   Line "线_136#mig1_2" at 219,318 size 114x103
      Visibility <- "ST_HMI_Var_HMI_r64Axis_ChengXing_Position_real2"
   Line "线_3" at 219,227 size 125x91
      Visibility <- "ST_HMI_Var_HMI_r64Axis_ChengXing_Position_real2"
   Line "线_4" at 219,273 size 149x45
      Visibility <- "ST_HMI_Var_HMI_r64Axis_ChengXing_Position_real2"
   Line "线_11#mig1_2" at 219,225 size 124x93
      Visibility <- "ST_HMI_Var_HMI_r64Axis_ChengXing_Position_real2"
   Line "线_5" at 219,276 size 150x41
      Visibility <- "ST_HMI_Var_HMI_r64Axis_ChengXing_Position_real2"
   Line "线_6" at 219,318 size 112x105
      Visibility <- "ST_HMI_Var_HMI_r64Axis_ChengXing_Position_real2"
   Line "线_157" at 219,229 size 126x88
      Visibility <- "ST_HMI_Var_HMI_r64Axis_ChengXing_Position_real2"
   Line "线_115#mig1_2" at 219,318 size 155x11
      Visibility <- "ST_HMI_Var_HMI_r64Axis_ChengXing_Position_real2"
   Line "线_7" at 219,318 size 143x61
      Visibility <- "ST_HMI_Var_HMI_r64Axis_ChengXing_Position_real2"
   Line "线_159" at 219,318 size 155x13
      Visibility <- "ST_HMI_Var_HMI_r64Axis_ChengXing_Position_real2"
   Line "线_8" at 219,318 size 141x63
      Visibility <- "ST_HMI_Var_HMI_r64Axis_ChengXing_Position_real2"
   Line "线_9" at 219,318 size 110x106
      Visibility <- "ST_HMI_Var_HMI_r64Axis_ChengXing_Position_real2"
   Line "线_13#mig1_2" at 219,231 size 127x87
      Visibility <- "ST_HMI_Var_HMI_r64Axis_ChengXing_Position_real2"
   Line "线_14" at 219,278 size 151x39
      Visibility <- "ST_HMI_Var_HMI_r64Axis_ChengXing_Position_real2"
   Line "线_22" at 219,318 size 155x15
      Visibility <- "ST_HMI_Var_HMI_r64Axis_ChengXing_Position_real2"
   Line "线_24" at 219,318 size 140x66
      Visibility <- "ST_HMI_Var_HMI_r64Axis_ChengXing_Position_real2"
   Line "线_25" at 219,318 size 108x108
      Visibility <- "ST_HMI_Var_HMI_r64Axis_ChengXing_Position_real2"
   Line "线_124#mig1_2" at 219,234 size 129x84
      Visibility <- "ST_HMI_Var_HMI_r64Axis_ChengXing_Position_real2"
   Line "线_27" at 219,282 size 151x36
      Visibility <- "ST_HMI_Var_HMI_r64Axis_ChengXing_Position_real2"
   Line "线_195" at 219,318 size 155x18
      Visibility <- "ST_HMI_Var_HMI_r64Axis_ChengXing_Position_real2"
   Line "线_196" at 219,318 size 139x69
      Visibility <- "ST_HMI_Var_HMI_r64Axis_ChengXing_Position_real2"
   Line "线_197" at 219,318 size 106x111
      Visibility <- "ST_HMI_Var_HMI_r64Axis_ChengXing_Position_real2"
   Line "线_198" at 219,236 size 131x81
      Visibility <- "ST_HMI_Var_HMI_r64Axis_ChengXing_Position_real2"
   Line "线_199" at 219,284 size 151x33
      Visibility <- "ST_HMI_Var_HMI_r64Axis_ChengXing_Position_real2"
   Line "线_200" at 219,318 size 154x21
      Visibility <- "ST_HMI_Var_HMI_r64Axis_ChengXing_Position_real2"
   Line "线_201" at 219,318 size 138x70
      Visibility <- "ST_HMI_Var_HMI_r64Axis_ChengXing_Position_real2"
   Line "线_202" at 219,318 size 104x112
      Visibility <- "ST_HMI_Var_HMI_r64Axis_ChengXing_Position_real2"
   Line "线_254" at 219,238 size 132x80
      Visibility <- "ST_HMI_Var_HMI_r64Axis_ChengXing_Position_real2"
   Line "线_255" at 219,287 size 152x31
      Visibility <- "ST_HMI_Var_HMI_r64Axis_ChengXing_Position_real2"
   Line "线_256" at 219,318 size 154x23
      Visibility <- "ST_HMI_Var_HMI_r64Axis_ChengXing_Position_real2"
   Line "线_257" at 219,318 size 136x73
      Visibility <- "ST_HMI_Var_HMI_r64Axis_ChengXing_Position_real2"
   Line "线_277" at 219,318 size 102x114
      Visibility <- "ST_HMI_Var_HMI_r64Axis_ChengXing_Position_real2"
   Line "线_278" at 219,240 size 133x77
      Visibility <- "ST_HMI_Var_HMI_r64Axis_ChengXing_Position_real2"
   Line "线_279" at 219,289 size 153x28
      Visibility <- "ST_HMI_Var_HMI_r64Axis_ChengXing_Position_real2"
   Line "线_280" at 219,318 size 153x27
      Visibility <- "ST_HMI_Var_HMI_r64Axis_ChengXing_Position_real2"
   Line "线_281" at 219,318 size 135x75
      Visibility <- "ST_HMI_Var_HMI_r64Axis_ChengXing_Position_real2"
   Line "线_282" at 219,318 size 100x116
      Visibility <- "ST_HMI_Var_HMI_r64Axis_ChengXing_Position_real2"
   Line "线_283" at 219,243 size 135x75
      Visibility <- "ST_HMI_Var_HMI_r64Axis_ChengXing_Position_real2"
   Line "线_125#mig1_2" at 219,291 size 153x27
      Visibility <- "ST_HMI_Var_HMI_r64Axis_ChengXing_Position_real2"
   Line "线_284" at 219,318 size 153x28
      Visibility <- "ST_HMI_Var_HMI_r64Axis_ChengXing_Position_real2"
   Line "线_285" at 219,318 size 133x77
      Visibility <- "ST_HMI_Var_HMI_r64Axis_ChengXing_Position_real2"
   Line "线_286" at 219,318 size 98x117
      Visibility <- "ST_HMI_Var_HMI_r64Axis_ChengXing_Position_real2"
   Line "线_287" at 219,245 size 136x73
      Visibility <- "ST_HMI_Var_HMI_r64Axis_ChengXing_Position_real2"
   Line "线_288" at 219,294 size 154x24
      Visibility <- "ST_HMI_Var_HMI_r64Axis_ChengXing_Position_real2"
   Line "线_289" at 219,318 size 152x32
      Visibility <- "ST_HMI_Var_HMI_r64Axis_ChengXing_Position_real2"
   Line "线_290" at 219,318 size 132x80
      Visibility <- "ST_HMI_Var_HMI_r64Axis_ChengXing_Position_real2"
   Line "线_291" at 219,318 size 96x119
      Visibility <- "ST_HMI_Var_HMI_r64Axis_ChengXing_Position_real2"
   Line "线_292" at 219,246 size 138x71
      Visibility <- "ST_HMI_Var_HMI_r64Axis_ChengXing_Position_real2"
   Line "线_293" at 219,296 size 155x21
      Visibility <- "ST_HMI_Var_HMI_r64Axis_ChengXing_Position_real2"
   Line "线_294" at 219,318 size 151x33
      Visibility <- "ST_HMI_Var_HMI_r64Axis_ChengXing_Position_real2"
   Line "线_295" at 219,318 size 131x82
      Visibility <- "ST_HMI_Var_HMI_r64Axis_ChengXing_Position_real2"
   Line "线_315" at 219,318 size 93x121
      Visibility <- "ST_HMI_Var_HMI_r64Axis_ChengXing_Position_real2"
   Line "线_316" at 219,249 size 139x69
      Visibility <- "ST_HMI_Var_HMI_r64Axis_ChengXing_Position_real2"
   Line "线_130#mig1_2" at 219,299 size 155x19
      Visibility <- "ST_HMI_Var_HMI_r64Axis_ChengXing_Position_real2"
   Line "线_317" at 219,318 size 92x123
      Visibility <- "ST_HMI_Var_HMI_r64Axis_ChengXing_Position_real2"
   Line "线_97#mig1_2" at 219,251 size 140x67
      Visibility <- "ST_HMI_Var_HMI_r64Axis_ChengXing_Position_real2"
   Line "线_129#mig1_2" at 219,301 size 155x16
      Visibility <- "ST_HMI_Var_HMI_r64Axis_ChengXing_Position_real2"
   Line "线_318" at 219,318 size 151x37
      Visibility <- "ST_HMI_Var_HMI_r64Axis_ChengXing_Position_real2"
   Line "线_319" at 219,318 size 129x84
      Visibility <- "ST_HMI_Var_HMI_r64Axis_ChengXing_Position_real2"
   Line "线_320" at 219,318 size 89x123
      Visibility <- "ST_HMI_Var_HMI_r64Axis_ChengXing_Position_real2"
   Line "线_321" at 219,253 size 141x64
      Visibility <- "ST_HMI_Var_HMI_r64Axis_ChengXing_Position_real2"
   Line "线_128#mig1_2" at 219,305 size 155x13
      Visibility <- "ST_HMI_Var_HMI_r64Axis_ChengXing_Position_real2"
   Line "线_322" at 219,318 size 151x39
      Visibility <- "ST_HMI_Var_HMI_r64Axis_ChengXing_Position_real2"
   Line "线_323" at 219,318 size 127x87
      Visibility <- "ST_HMI_Var_HMI_r64Axis_ChengXing_Position_real2"
   Line "线_324" at 219,256 size 143x62
      Visibility <- "ST_HMI_Var_HMI_r64Axis_ChengXing_Position_real2"
   Line "线_131#mig1_2" at 219,306 size 155x11
      Visibility <- "ST_HMI_Var_HMI_r64Axis_ChengXing_Position_real2"
   Line "线_325" at 219,318 size 150x42
      Visibility <- "ST_HMI_Var_HMI_r64Axis_ChengXing_Position_real2"
   Line "线_326" at 219,318 size 126x89
      Visibility <- "ST_HMI_Var_HMI_r64Axis_ChengXing_Position_real2"
   Line "线_114#mig1_2" at 219,258 size 144x59
      Visibility <- "ST_HMI_Var_HMI_r64Axis_ChengXing_Position_real2"
   Line "线_327" at 219,310 size 156x8
      Visibility <- "ST_HMI_Var_HMI_r64Axis_ChengXing_Position_real2"
   Line "线_328" at 219,318 size 149x45
      Visibility <- "ST_HMI_Var_HMI_r64Axis_ChengXing_Position_real2"
   Line "线_329" at 219,318 size 125x91
      Visibility <- "ST_HMI_Var_HMI_r64Axis_ChengXing_Position_real2"
   Line "线_120#mig1_2" at 219,261 size 144x57
      Visibility <- "ST_HMI_Var_HMI_r64Axis_ChengXing_Position_real2"
   Line "线_330" at 219,312 size 156x5
      Visibility <- "ST_HMI_Var_HMI_r64Axis_ChengXing_Position_real2"
   Line "线_331" at 219,318 size 148x47
      Visibility <- "ST_HMI_Var_HMI_r64Axis_ChengXing_Position_real2"
   Line "线_332" at 219,318 size 123x93
      Visibility <- "ST_HMI_Var_HMI_r64Axis_ChengXing_Position_real2"
   Line "线_333" at 219,264 size 145x54
      Visibility <- "ST_HMI_Var_HMI_r64Axis_ChengXing_Position_real2"
   Line "线_150#mig1_2" at 219,315 size 156x3
      Visibility <- "ST_HMI_Var_HMI_r64Axis_ChengXing_Position_real2"
   Line "线_334" at 219,318 size 147x50
      Visibility <- "ST_HMI_Var_HMI_r64Axis_ChengXing_Position_real2"
   Line "线_335" at 219,318 size 121x95
      Visibility <- "ST_HMI_Var_HMI_r64Axis_ChengXing_Position_real2"
   Line "线_336" at 219,266 size 146x51
      Visibility <- "ST_HMI_Var_HMI_r64Axis_ChengXing_Position_real2"
   Line "线_147#mig1_2" at 219,318 size 156x0
      Visibility <- "ST_HMI_Var_HMI_r64Axis_ChengXing_Position_real2"
   Line "线_337" at 219,318 size 146x52
      Visibility <- "ST_HMI_Var_HMI_r64Axis_ChengXing_Position_real2"
   Line "线_338" at 219,318 size 119x98
      Visibility <- "ST_HMI_Var_HMI_r64Axis_ChengXing_Position_real2"
   Line "线_339" at 219,268 size 147x50
      Visibility <- "ST_HMI_Var_HMI_r64Axis_ChengXing_Position_real2"
   Line "线_340" at 219,318 size 156x3
      Visibility <- "ST_HMI_Var_HMI_r64Axis_ChengXing_Position_real2"
   Line "线_341" at 219,318 size 145x54
      Visibility <- "ST_HMI_Var_HMI_r64Axis_ChengXing_Position_real2"
   Line "线_342" at 219,318 size 144x57
      Visibility <- "ST_HMI_Var_HMI_r64Axis_ChengXing_Position_real2"
   Line "线_343" at 219,318 size 118x99
      Visibility <- "ST_HMI_Var_HMI_r64Axis_ChengXing_Position_real2"
   Line "线_344" at 219,318 size 116x101
      Visibility <- "ST_HMI_Var_HMI_r64Axis_ChengXing_Position_real2"
   Line "线_345" at 219,271 size 148x46
      Visibility <- "ST_HMI_Var_HMI_r64Axis_ChengXing_Position_real2"
   Line "线_346" at 219,318 size 156x5
      Visibility <- "ST_HMI_Var_HMI_r64Axis_ChengXing_Position_real2"
   Line "线_29" at 219,318 size 156x8
      Visibility <- "ST_HMI_Var_HMI_r64Axis_ChengXing_Position_real2"
   Line "线_31" at 219,318 size 144x58
      Visibility <- "ST_HMI_Var_HMI_r64Axis_ChengXing_Position_real2"
   Line "线_136#mig1_1" at 219,318 size 114x103
      Visibility <- "ST_HMI_Var_HMI_r64Axis_ChengXing_Position_real2"
   Line "线_38" at 219,227 size 125x91
      Visibility <- "ST_HMI_Var_HMI_r64Axis_ChengXing_Position_real2"
   Line "线_39" at 219,273 size 149x45
      Visibility <- "ST_HMI_Var_HMI_r64Axis_ChengXing_Position_real2"
   Line "线_11#mig1_1" at 219,225 size 124x93
      Visibility <- "ST_HMI_Var_HMI_r64Axis_ChengXing_Position_real2"
   Line "线_41" at 219,276 size 150x41
      Visibility <- "ST_HMI_Var_HMI_r64Axis_ChengXing_Position_real2"
   Line "线_43" at 219,318 size 112x105
      Visibility <- "ST_HMI_Var_HMI_r64Axis_ChengXing_Position_real2"
   Line "线_44" at 219,229 size 126x88
      Visibility <- "ST_HMI_Var_HMI_r64Axis_ChengXing_Position_real2"
   Line "线_115#mig1_1" at 219,318 size 155x11
      Visibility <- "ST_HMI_Var_HMI_r64Axis_ChengXing_Position_real2"
   Line "线_46" at 219,318 size 143x61
      Visibility <- "ST_HMI_Var_HMI_r64Axis_ChengXing_Position_real2"
   Line "线_47" at 219,318 size 155x13
      Visibility <- "ST_HMI_Var_HMI_r64Axis_ChengXing_Position_real2"
   Line "线_48" at 219,318 size 141x63
      Visibility <- "ST_HMI_Var_HMI_r64Axis_ChengXing_Position_real2"
   Line "线_49" at 219,318 size 110x106
      Visibility <- "ST_HMI_Var_HMI_r64Axis_ChengXing_Position_real2"
   Line "线_13#mig1_1" at 219,231 size 127x87
      Visibility <- "ST_HMI_Var_HMI_r64Axis_ChengXing_Position_real2"
   Line "线_59" at 219,278 size 151x39
      Visibility <- "ST_HMI_Var_HMI_r64Axis_ChengXing_Position_real2"
   Line "线_60" at 219,318 size 155x15
      Visibility <- "ST_HMI_Var_HMI_r64Axis_ChengXing_Position_real2"
   Line "线_61" at 219,318 size 140x66
      Visibility <- "ST_HMI_Var_HMI_r64Axis_ChengXing_Position_real2"
   Line "线_65" at 219,318 size 108x108
      Visibility <- "ST_HMI_Var_HMI_r64Axis_ChengXing_Position_real2"
   Line "线_124#mig1_1" at 219,234 size 129x84
      Visibility <- "ST_HMI_Var_HMI_r64Axis_ChengXing_Position_real2"
   Line "线_66" at 219,282 size 151x36
      Visibility <- "ST_HMI_Var_HMI_r64Axis_ChengXing_Position_real2"
   Line "线_67" at 219,318 size 155x18
      Visibility <- "ST_HMI_Var_HMI_r64Axis_ChengXing_Position_real2"
   Line "线_69" at 219,318 size 139x69
      Visibility <- "ST_HMI_Var_HMI_r64Axis_ChengXing_Position_real2"
   Line "线_70" at 219,318 size 106x111
      Visibility <- "ST_HMI_Var_HMI_r64Axis_ChengXing_Position_real2"
   Line "线_71" at 219,236 size 131x81
      Visibility <- "ST_HMI_Var_HMI_r64Axis_ChengXing_Position_real2"
   Line "线_72" at 219,284 size 151x33
      Visibility <- "ST_HMI_Var_HMI_r64Axis_ChengXing_Position_real2"
   Line "线_73" at 219,318 size 154x21
      Visibility <- "ST_HMI_Var_HMI_r64Axis_ChengXing_Position_real2"
   Line "线_74" at 219,318 size 138x70
      Visibility <- "ST_HMI_Var_HMI_r64Axis_ChengXing_Position_real2"
   Line "线_76" at 219,318 size 104x112
      Visibility <- "ST_HMI_Var_HMI_r64Axis_ChengXing_Position_real2"
   Line "线_77" at 219,238 size 132x80
      Visibility <- "ST_HMI_Var_HMI_r64Axis_ChengXing_Position_real2"
   Line "线_78" at 219,287 size 152x31
      Visibility <- "ST_HMI_Var_HMI_r64Axis_ChengXing_Position_real2"
   Line "线_79" at 219,318 size 154x23
      Visibility <- "ST_HMI_Var_HMI_r64Axis_ChengXing_Position_real2"
   Line "线_82" at 219,318 size 136x73
      Visibility <- "ST_HMI_Var_HMI_r64Axis_ChengXing_Position_real2"
   Line "线_84" at 219,318 size 102x114
      Visibility <- "ST_HMI_Var_HMI_r64Axis_ChengXing_Position_real2"
   Line "线_86" at 219,240 size 133x77
      Visibility <- "ST_HMI_Var_HMI_r64Axis_ChengXing_Position_real2"
   Line "线_87" at 219,289 size 153x28
      Visibility <- "ST_HMI_Var_HMI_r64Axis_ChengXing_Position_real2"
   Line "线_88" at 219,318 size 153x27
      Visibility <- "ST_HMI_Var_HMI_r64Axis_ChengXing_Position_real2"
   Line "线_90" at 219,318 size 135x75
      Visibility <- "ST_HMI_Var_HMI_r64Axis_ChengXing_Position_real2"
   Line "线_92" at 219,318 size 100x116
      Visibility <- "ST_HMI_Var_HMI_r64Axis_ChengXing_Position_real2"
   Line "线_93" at 219,243 size 135x75
      Visibility <- "ST_HMI_Var_HMI_r64Axis_ChengXing_Position_real2"
   Line "线_125#mig1_1" at 219,291 size 153x27
      Visibility <- "ST_HMI_Var_HMI_r64Axis_ChengXing_Position_real2"
   Line "线_98" at 219,318 size 153x28
      Visibility <- "ST_HMI_Var_HMI_r64Axis_ChengXing_Position_real2"
   Line "线_99" at 219,318 size 133x77
      Visibility <- "ST_HMI_Var_HMI_r64Axis_ChengXing_Position_real2"
   Line "线_109" at 219,318 size 98x117
      Visibility <- "ST_HMI_Var_HMI_r64Axis_ChengXing_Position_real2"
   Line "线_117" at 219,245 size 136x73
      Visibility <- "ST_HMI_Var_HMI_r64Axis_ChengXing_Position_real2"
   Line "线_119" at 219,294 size 154x24
      Visibility <- "ST_HMI_Var_HMI_r64Axis_ChengXing_Position_real2"
   Line "线_132" at 219,318 size 152x32
      Visibility <- "ST_HMI_Var_HMI_r64Axis_ChengXing_Position_real2"
   Line "线_135" at 219,318 size 132x80
      Visibility <- "ST_HMI_Var_HMI_r64Axis_ChengXing_Position_real2"
   Line "线_138" at 219,318 size 96x119
      Visibility <- "ST_HMI_Var_HMI_r64Axis_ChengXing_Position_real2"
   Line "线_347" at 219,246 size 138x71
      Visibility <- "ST_HMI_Var_HMI_r64Axis_ChengXing_Position_real2"
   Line "线_348" at 219,296 size 155x21
      Visibility <- "ST_HMI_Var_HMI_r64Axis_ChengXing_Position_real2"
   Line "线_349" at 219,318 size 151x33
      Visibility <- "ST_HMI_Var_HMI_r64Axis_ChengXing_Position_real2"
   Line "线_350" at 219,318 size 131x82
      Visibility <- "ST_HMI_Var_HMI_r64Axis_ChengXing_Position_real2"
   Line "线_351" at 219,318 size 93x121
      Visibility <- "ST_HMI_Var_HMI_r64Axis_ChengXing_Position_real2"
   Line "线_352" at 219,249 size 139x69
      Visibility <- "ST_HMI_Var_HMI_r64Axis_ChengXing_Position_real2"
   Line "线_130#mig1_1" at 219,299 size 155x19
      Visibility <- "ST_HMI_Var_HMI_r64Axis_ChengXing_Position_real2"
   Line "线_353" at 219,318 size 92x123
      Visibility <- "ST_HMI_Var_HMI_r64Axis_ChengXing_Position_real2"
   Line "线_97#mig1_1" at 219,251 size 140x67
      Visibility <- "ST_HMI_Var_HMI_r64Axis_ChengXing_Position_real2"
   Line "线_129#mig1_1" at 219,301 size 155x16
      Visibility <- "ST_HMI_Var_HMI_r64Axis_ChengXing_Position_real2"
   Line "线_354" at 219,318 size 151x37
      Visibility <- "ST_HMI_Var_HMI_r64Axis_ChengXing_Position_real2"
   Line "线_355" at 219,318 size 129x84
      Visibility <- "ST_HMI_Var_HMI_r64Axis_ChengXing_Position_real2"
   Line "线_356" at 219,318 size 89x123
      Visibility <- "ST_HMI_Var_HMI_r64Axis_ChengXing_Position_real2"
   Line "线_357" at 219,253 size 141x64
      Visibility <- "ST_HMI_Var_HMI_r64Axis_ChengXing_Position_real2"
   Line "线_128#mig1_1" at 219,305 size 155x13
      Visibility <- "ST_HMI_Var_HMI_r64Axis_ChengXing_Position_real2"
   Line "线_358" at 219,318 size 151x39
      Visibility <- "ST_HMI_Var_HMI_r64Axis_ChengXing_Position_real2"
   Line "线_359" at 219,318 size 127x87
      Visibility <- "ST_HMI_Var_HMI_r64Axis_ChengXing_Position_real2"
   Line "线_360" at 219,256 size 143x62
      Visibility <- "ST_HMI_Var_HMI_r64Axis_ChengXing_Position_real2"
   Line "线_131#mig1_1" at 219,306 size 155x11
      Visibility <- "ST_HMI_Var_HMI_r64Axis_ChengXing_Position_real2"
   Line "线_361" at 219,318 size 150x42
      Visibility <- "ST_HMI_Var_HMI_r64Axis_ChengXing_Position_real2"
   Line "线_362" at 219,318 size 126x89
      Visibility <- "ST_HMI_Var_HMI_r64Axis_ChengXing_Position_real2"
   Line "线_114#mig1_1" at 219,258 size 144x59
      Visibility <- "ST_HMI_Var_HMI_r64Axis_ChengXing_Position_real2"
   Line "线_363" at 219,310 size 156x8
      Visibility <- "ST_HMI_Var_HMI_r64Axis_ChengXing_Position_real2"
   Line "线_364" at 219,318 size 149x45
      Visibility <- "ST_HMI_Var_HMI_r64Axis_ChengXing_Position_real2"
   Line "线_365" at 219,318 size 125x91
      Visibility <- "ST_HMI_Var_HMI_r64Axis_ChengXing_Position_real2"
   Line "线_120#mig1_1" at 219,261 size 144x57
      Visibility <- "ST_HMI_Var_HMI_r64Axis_ChengXing_Position_real2"
   Line "线_366" at 219,312 size 156x5
      Visibility <- "ST_HMI_Var_HMI_r64Axis_ChengXing_Position_real2"
   Line "线_367" at 219,318 size 148x47
      Visibility <- "ST_HMI_Var_HMI_r64Axis_ChengXing_Position_real2"
   Line "线_368" at 219,318 size 123x93
      Visibility <- "ST_HMI_Var_HMI_r64Axis_ChengXing_Position_real2"
   Line "线_369" at 219,264 size 145x54
      Visibility <- "ST_HMI_Var_HMI_r64Axis_ChengXing_Position_real2"
   Line "线_150#mig1_1" at 219,315 size 156x3
      Visibility <- "ST_HMI_Var_HMI_r64Axis_ChengXing_Position_real2"
   Line "线_370" at 219,318 size 147x50
      Visibility <- "ST_HMI_Var_HMI_r64Axis_ChengXing_Position_real2"
   Line "线_371" at 219,318 size 121x95
      Visibility <- "ST_HMI_Var_HMI_r64Axis_ChengXing_Position_real2"
   Line "线_372" at 219,266 size 146x51
      Visibility <- "ST_HMI_Var_HMI_r64Axis_ChengXing_Position_real2"
   Line "线_147#mig1_1" at 219,318 size 156x0
      Visibility <- "ST_HMI_Var_HMI_r64Axis_ChengXing_Position_real2"
   Line "线_373" at 219,318 size 146x52
      Visibility <- "ST_HMI_Var_HMI_r64Axis_ChengXing_Position_real2"
   Line "线_374" at 219,318 size 119x98
      Visibility <- "ST_HMI_Var_HMI_r64Axis_ChengXing_Position_real2"
   Line "线_375" at 219,268 size 147x50
      Visibility <- "ST_HMI_Var_HMI_r64Axis_ChengXing_Position_real2"
   Line "线_376" at 219,318 size 156x3
      Visibility <- "ST_HMI_Var_HMI_r64Axis_ChengXing_Position_real2"
   Line "线_377" at 219,318 size 145x54
      Visibility <- "ST_HMI_Var_HMI_r64Axis_ChengXing_Position_real2"
   Line "线_378" at 219,318 size 144x57
      Visibility <- "ST_HMI_Var_HMI_r64Axis_ChengXing_Position_real2"
   Line "线_379" at 219,318 size 118x99
      Visibility <- "ST_HMI_Var_HMI_r64Axis_ChengXing_Position_real2"
   Line "线_380" at 219,318 size 116x101
      Visibility <- "ST_HMI_Var_HMI_r64Axis_ChengXing_Position_real2"
   Line "线_381" at 219,271 size 148x46
      Visibility <- "ST_HMI_Var_HMI_r64Axis_ChengXing_Position_real2"
   Line "线_382" at 219,318 size 156x5
      Visibility <- "ST_HMI_Var_HMI_r64Axis_ChengXing_Position_real2"
   Polygon "多边形_8" at 292,385 size 21x46
      Visibility <- "VBS_hengsi_status0"
   Polygon "多边形_7" at 288,376 size 31x55
      Visibility <- "VBS_hengsi_status0"
   Polygon "多边形_10" at 287,367 size 36x63
      Visibility <- "VBS_hengsi_status0"
   Polygon "多边形_11#mig1" at 287,361 size 40x70
      Visibility <- "VBS_hengsi_status0"
   Polygon "多边形_12" at 285,354 size 45x77
      Visibility <- "VBS_hengsi_status0"
   Polygon "多边形_18" at 285,345 size 45x86
      Visibility <- "VBS_hengsi_status1"
   Polygon "多边形_17" at 285,338 size 49x93
      Visibility <- "VBS_hengsi_status1"
   Polygon "多边形_16" at 287,328 size 50x103
      Visibility <- "VBS_hengsi_status1"
   Polygon "多边形_15" at 287,318 size 54x115
      Visibility <- "VBS_hengsi_status1"
   Polygon "多边形_14" at 287,309 size 56x123
      Visibility <- "VBS_hengsi_status1"
   Polygon "多边形_19" at 285,301 size 59x132
      Visibility <- "VBS_hengsi_status1"
   Polygon "多边形_20" at 287,289 size 61x144
      Visibility <- "VBS_hengsi_status1"
   Polygon "多边形_21" at 285,283 size 64x149
      Visibility <- "VBS_hengsi_status1"
   Polygon "多边形_22" at 285,278 size 66x154
      Visibility <- "VBS_hengsi_status1"
   Group "Group_9" at 162,225 size 228x110
   Group "Group_10" at 162,225 size 228x110
   Line "线_10" at 188,297 size 202x7
      Visibility <- "ST_HMI_Var_HMI_r64Axis_1_ZhangLi_Position_JuanRao_real2"
   Line "线_12" at 188,305 size 202x0
      Visibility <- "ST_HMI_Var_HMI_r64Axis_1_ZhangLi_Position_JuanRao_real2"
   Line "线_17" at 188,301 size 202x4
      Visibility <- "ST_HMI_Var_HMI_r64Axis_1_ZhangLi_Position_JuanRao_real2"
   Line "线_18" at 188,305 size 202x4
      Visibility <- "ST_HMI_Var_HMI_r64Axis_1_ZhangLi_Position_JuanRao_real2"
   Line "线_19" at 188,305 size 202x7
      Visibility <- "ST_HMI_Var_HMI_r64Axis_1_ZhangLi_Position_JuanRao_real2"
   Line "线_20" at 188,305 size 202x11
      Visibility <- "ST_HMI_Var_HMI_r64Axis_1_ZhangLi_Position_JuanRao_real2"
   Line "线_116" at 188,305 size 201x15
      Visibility <- "ST_HMI_Var_HMI_r64Axis_1_ZhangLi_Position_JuanRao_real2"
   Line "线_118" at 188,305 size 201x19
      Visibility <- "ST_HMI_Var_HMI_r64Axis_1_ZhangLi_Position_JuanRao_real2"
   Line "线_121" at 188,305 size 201x23
      Visibility <- "ST_HMI_Var_HMI_r64Axis_1_ZhangLi_Position_JuanRao_real2"
   Line "线_126" at 188,305 size 200x27
      Visibility <- "ST_HMI_Var_HMI_r64Axis_1_ZhangLi_Position_JuanRao_real2"
   Line "线_127" at 188,305 size 200x30
      Visibility <- "ST_HMI_Var_HMI_r64Axis_1_ZhangLi_Position_JuanRao_real2"
   Line "线_128" at 188,225 size 187x80
      Visibility <- "ST_HMI_Var_HMI_r64Axis_1_ZhangLi_Position_JuanRao_real2"
   Line "线_129" at 188,229 size 189x76
      Visibility <- "ST_HMI_Var_HMI_r64Axis_1_ZhangLi_Position_JuanRao_real2"
   Line "线_130" at 188,231 size 190x73
      Visibility <- "ST_HMI_Var_HMI_r64Axis_1_ZhangLi_Position_JuanRao_real2"
   Line "线_131" at 188,235 size 191x70
      Visibility <- "ST_HMI_Var_HMI_r64Axis_1_ZhangLi_Position_JuanRao_real2"
   Line "线_133" at 188,239 size 192x66
      Visibility <- "ST_HMI_Var_HMI_r64Axis_1_ZhangLi_Position_JuanRao_real2"
   Line "线_134" at 188,242 size 193x62
      Visibility <- "ST_HMI_Var_HMI_r64Axis_1_ZhangLi_Position_JuanRao_real2"
   Line "线_136" at 188,246 size 194x59
      Visibility <- "ST_HMI_Var_HMI_r64Axis_1_ZhangLi_Position_JuanRao_real2"
   Line "线_137" at 188,250 size 195x55
      Visibility <- "ST_HMI_Var_HMI_r64Axis_1_ZhangLi_Position_JuanRao_real2"
   Line "线_139" at 188,253 size 196x51
      Visibility <- "ST_HMI_Var_HMI_r64Axis_1_ZhangLi_Position_JuanRao_real2"
   Line "线_140" at 188,257 size 197x48
      Visibility <- "ST_HMI_Var_HMI_r64Axis_1_ZhangLi_Position_JuanRao_real2"
   Line "线_141" at 188,261 size 198x44
      Visibility <- "ST_HMI_Var_HMI_r64Axis_1_ZhangLi_Position_JuanRao_real2"
   Line "线_142" at 188,264 size 199x40
      Visibility <- "ST_HMI_Var_HMI_r64Axis_1_ZhangLi_Position_JuanRao_real2"
   Line "线_143" at 188,268 size 199x37
      Visibility <- "ST_HMI_Var_HMI_r64Axis_1_ZhangLi_Position_JuanRao_real2"
   Line "线_144" at 188,272 size 199x33
      Visibility <- "ST_HMI_Var_HMI_r64Axis_1_ZhangLi_Position_JuanRao_real2"
   Line "线_145" at 188,275 size 200x29
      Visibility <- "ST_HMI_Var_HMI_r64Axis_1_ZhangLi_Position_JuanRao_real2"
   Line "线_146" at 188,279 size 200x26
      Visibility <- "ST_HMI_Var_HMI_r64Axis_1_ZhangLi_Position_JuanRao_real2"
   Line "线_147" at 188,283 size 201x22
      Visibility <- "ST_HMI_Var_HMI_r64Axis_1_ZhangLi_Position_JuanRao_real2"
   Line "线_148" at 188,285 size 201x19
      Visibility <- "ST_HMI_Var_HMI_r64Axis_1_ZhangLi_Position_JuanRao_real2"
   Line "线_149" at 188,290 size 201x15
      Visibility <- "ST_HMI_Var_HMI_r64Axis_1_ZhangLi_Position_JuanRao_real2"
   Line "线_150" at 188,294 size 202x11
      Visibility <- "ST_HMI_Var_HMI_r64Axis_1_ZhangLi_Position_JuanRao_real2"
   Line "线_151" at 188,297 size 202x7
      Visibility <- "ST_HMI_Var_HMI_r64Axis_1_ZhangLi_Position_JuanRao_real2"
   Line "线_152" at 188,305 size 202x0
      Visibility <- "ST_HMI_Var_HMI_r64Axis_1_ZhangLi_Position_JuanRao_real2"
   Line "线_153" at 188,301 size 202x4
      Visibility <- "ST_HMI_Var_HMI_r64Axis_1_ZhangLi_Position_JuanRao_real2"
   Line "线_154" at 188,305 size 202x4
      Visibility <- "ST_HMI_Var_HMI_r64Axis_1_ZhangLi_Position_JuanRao_real2"
   Line "线_155" at 188,305 size 202x7
      Visibility <- "ST_HMI_Var_HMI_r64Axis_1_ZhangLi_Position_JuanRao_real2"
   Line "线_156" at 188,305 size 202x11
      Visibility <- "ST_HMI_Var_HMI_r64Axis_1_ZhangLi_Position_JuanRao_real2"
   Line "线_158" at 188,305 size 201x15
      Visibility <- "ST_HMI_Var_HMI_r64Axis_1_ZhangLi_Position_JuanRao_real2"
   Line "线_160" at 188,305 size 201x19
      Visibility <- "ST_HMI_Var_HMI_r64Axis_1_ZhangLi_Position_JuanRao_real2"
   Line "线_161" at 188,305 size 201x23
      Visibility <- "ST_HMI_Var_HMI_r64Axis_1_ZhangLi_Position_JuanRao_real2"
   Line "线_162" at 188,305 size 200x27
      Visibility <- "ST_HMI_Var_HMI_r64Axis_1_ZhangLi_Position_JuanRao_real2"
   Line "线_163" at 188,305 size 200x30
      Visibility <- "ST_HMI_Var_HMI_r64Axis_1_ZhangLi_Position_JuanRao_real2"
   Line "线_164" at 188,225 size 187x80
      Visibility <- "ST_HMI_Var_HMI_r64Axis_1_ZhangLi_Position_JuanRao_real2"
   Line "线_165" at 188,229 size 189x76
      Visibility <- "ST_HMI_Var_HMI_r64Axis_1_ZhangLi_Position_JuanRao_real2"
   Line "线_166" at 188,231 size 190x73
      Visibility <- "ST_HMI_Var_HMI_r64Axis_1_ZhangLi_Position_JuanRao_real2"
   Line "线_167" at 188,235 size 191x70
      Visibility <- "ST_HMI_Var_HMI_r64Axis_1_ZhangLi_Position_JuanRao_real2"
   Line "线_168" at 188,239 size 192x66
      Visibility <- "ST_HMI_Var_HMI_r64Axis_1_ZhangLi_Position_JuanRao_real2"
   Line "线_169" at 188,242 size 193x62
      Visibility <- "ST_HMI_Var_HMI_r64Axis_1_ZhangLi_Position_JuanRao_real2"
   Line "线_170" at 188,246 size 194x59
      Visibility <- "ST_HMI_Var_HMI_r64Axis_1_ZhangLi_Position_JuanRao_real2"
   Line "线_171" at 188,250 size 195x55
      Visibility <- "ST_HMI_Var_HMI_r64Axis_1_ZhangLi_Position_JuanRao_real2"
   Line "线_172" at 188,253 size 196x51
      Visibility <- "ST_HMI_Var_HMI_r64Axis_1_ZhangLi_Position_JuanRao_real2"
   Line "线_173" at 188,257 size 197x48
      Visibility <- "ST_HMI_Var_HMI_r64Axis_1_ZhangLi_Position_JuanRao_real2"
   Line "线_174" at 188,261 size 198x44
      Visibility <- "ST_HMI_Var_HMI_r64Axis_1_ZhangLi_Position_JuanRao_real2"
   Line "线_175" at 188,264 size 199x40
      Visibility <- "ST_HMI_Var_HMI_r64Axis_1_ZhangLi_Position_JuanRao_real2"
   Line "线_176" at 188,268 size 199x37
      Visibility <- "ST_HMI_Var_HMI_r64Axis_1_ZhangLi_Position_JuanRao_real2"
   Line "线_177" at 188,272 size 199x33
      Visibility <- "ST_HMI_Var_HMI_r64Axis_1_ZhangLi_Position_JuanRao_real2"
   Line "线_178" at 188,275 size 200x29
      Visibility <- "ST_HMI_Var_HMI_r64Axis_1_ZhangLi_Position_JuanRao_real2"
   Line "线_179" at 188,279 size 200x26
      Visibility <- "ST_HMI_Var_HMI_r64Axis_1_ZhangLi_Position_JuanRao_real2"
   Line "线_180" at 188,283 size 201x22
      Visibility <- "ST_HMI_Var_HMI_r64Axis_1_ZhangLi_Position_JuanRao_real2"
   Line "线_181" at 188,285 size 201x19
      Visibility <- "ST_HMI_Var_HMI_r64Axis_1_ZhangLi_Position_JuanRao_real2"
   Line "线_182" at 188,290 size 201x15
      Visibility <- "ST_HMI_Var_HMI_r64Axis_1_ZhangLi_Position_JuanRao_real2"
   Line "线_183" at 188,294 size 202x11
      Visibility <- "ST_HMI_Var_HMI_r64Axis_1_ZhangLi_Position_JuanRao_real2"
   TextField "文本域_2" at 1139,375 size 32x36; Text 'mm'
   IOField "IO Field_1" at 1053,375 size 86x39; FormatPattern 9999.9
      ProcessValue <- "ST_HMI_Var_HMI_r64_ZouChe_ZhanJu_Max_Effect"
   TextField "文本域_1" at 556,323 size 22x25; Text 'mm'
   IOField "IO Field_51" at 420,323 size 60x25; FormatPattern 9999.9
      ProcessValue <- "ST_HMI_Var_HMI_r64Axis_ZouChe_Position_real"
   IOField "IO Field_2" at 496,323 size 60x25; FormatPattern 9999.9
      ProcessValue <- "ST_HMI_Var_HMI_r64Axis_ZouChe_Position_object"
   TextField "文本域_3" at 480,323 size 16x25; Text '/'
   TextField "文本域_12" at 163,221 size 41x24; Text '张力'
   IOField "IO Field_74" at 202,245 size 51x24; FormatPattern 999.9
      ProcessValue <- "ST_HMI_Var_HMI_r64Axis_ChengXing_Position_real"
   TextField "文本域_11" at 163,245 size 41x24; Text '成形'
   IOField "IO Field_80" at 202,221 size 51x24; FormatPattern 999.9
      ProcessValue <- "ST_HMI_Var_HMI_r64Axis_1_ZhangLi_Position_JuanRao_real"
   IOField "IO Field_3" at 163,155 size 42x25; FormatPattern 9999
      Visibility <- "ST_Main_Var_g_i16_Mode_Enabled"
      ProcessValue <- "ST_HMI_Var_HMI_r64NianDu_real_ShengTou"
   IOField "IO Field_53" at 163,180 size 42x25; FormatPattern 9999
      ProcessValue <- "ST_HMI_Var_HMI_r64Niandu_all_Current"
   TextField "文本域_6" at 205,155 size 56x25; Text '/'
   IOField "IO Field_54" at 163,155 size 42x25; FormatPattern 9999
      Visibility <- "ST_Main_Var_g_i16_Mode_Enabled"
      ProcessValue <- "ST_HMI_Var_HMI_r64NianDu_real"
   TextField "文本域_7" at 205,180 size 56x25; Text '捻/米'

Template "模板_调试" 1280x740
   Button "template_test_1" at 80,680 size 80x60; TextOn '手动画面'; TextOff '手动操作'; PictureOn "manual_5_500×500_反相"; PictureOff "manual_5_500×500"
      on Release: ActivateScreenByNumber("Picture", 0)
      on Press: SetTag("Picture", 5)
      Appearance <- "Picture"
   Button "template_test_2" at 720,680 size 80x60; TextOn '报警画面'; TextOff '报 警'; PictureOn "emblem_important_1_200×200_反相"; PictureOff "emblem_important_1_200×200"
      on Release: ActivateScreenByNumber("Picture", 0)
      on Press: SetTag("Picture", 6)
      Appearance <- "Picture"
   Button "template_test_5" at 800,680 size 80x60; TextOn '保养提示'; TextOff '保养提示'; PictureOn "baoyang_6_600×600_反相"; PictureOff "baoyang_6_600×600"
      on Release: ActivateScreenByNumber("Picture", 0)
      on Press: SetTag("Picture", 8)
      Appearance <- "Picture"
   Button "template_test_7" at 880,680 size 80x60; TextOn '调试画面'; TextOff '调 试'; Authorization "Operate_4"; PictureOff "kdeconnect-tray_100×100"; PictureOn "kdeconnect-tray_100×100_反相"
      on Release: ActivateScreenByNumber("Picture", 0); function_f23ef4c9()
      on Press: SetTag("Picture", 3)
      Appearance <- "Picture"
   Button "template_test_3" at 0,680 size 80x60; TextOn '手动画面'; TextOff '手动操作'; PictureOff "图形_16"
      on Release: ActivateScreenByNumber("Picture", 0); SetTag("ST_HMI_Var_HMI_i32_ZouChe_ZhanJu_ss_1", 0)
      on Press: function_f23ef4c9(); SetTag("Picture", 1)
      Appearance <- "Picture"
   Button "template_test_4" at 1120,680 size 80x60; TextOff '调 试'; TextOn '调试画面'; PictureOn "System_Shutdown_反相_100×100"; PictureOff "System_Shutdown_100×100"; Authorization "Operate_4"
      on Click: function_f23ef4c9()
      on Release: StopRuntime(0)
   Button "template_test_6" at 1040,680 size 80x60; TextOff 'Text'; TextOn '调试画面'; PictureOn "computer_laptop_100×100_反相"; PictureOff "computer_laptop_100×100"; Authorization "Operate_4"
      on Click: function_f23ef4c9()
      on Release: function_f34a74f3()
   Button "template_test_8" at 960,680 size 80x60; TextOff 'Text'; TextOn '调试画面'; PictureOn "similarartists_amarok_100×100_反相"; PictureOff "similarartists_amarok_100×100"; Authorization "Operate_4"
      on Release: ActivateScreenByNumber("Picture", 0); function_f23ef4c9()
      on Press: SetTag("Picture", 7)
      Appearance <- "Picture"
   Button "template_test_9" at 0,20 size 130x47; TextOn '1牵伸相关'; TextOff '1牵伸相关'
      on Release: ActivateScreenByNumber("Picture", 0); SetTag("ST_HMI_Var_HMI_i32_ZouChe_ZhanJu_ss_1", 0)
      on Press: SetTag("Picture", 31)
      Appearance <- "Picture"
   Button "template_test_10" at 0,85 size 130x47; TextOn '2加捻相关'; TextOff '2加捻相关'
      on Release: ActivateScreenByNumber("Picture", 0); SetTag("ST_HMI_Var_HMI_i32_ZouChe_ZhanJu_ss_1", 0)
      on Press: SetTag("Picture", 32)
      Appearance <- "Picture"
   Button "template_test_11" at 0,151 size 130x47; TextOn '3退绕相关1'; TextOff '3退绕相关1'
      on Release: ActivateScreenByNumber("Picture", 0); SetTag("ST_HMI_Var_HMI_i32_ZouChe_ZhanJu_ss_1", 0)
      on Press: SetTag("Picture", 33)
      Appearance <- "Picture"
   Button "template_test_12" at 0,216 size 130x47; TextOn '4退绕相关2'; TextOff '4退绕相关2'
      on Release: ActivateScreenByNumber("Picture", 0); SetTag("ST_HMI_Var_HMI_i32_ZouChe_ZhanJu_ss_1", 0)
      on Press: SetTag("Picture", 34)
      Appearance <- "Picture"
   Button "template_test_13" at 0,282 size 130x47; TextOn '5成形相关'; TextOff '5成形相关'
      on Release: ActivateScreenByNumber("Picture", 0); SetTag("ST_HMI_Var_HMI_i32_ZouChe_ZhanJu_ss_1", 0)
      on Press: SetTag("Picture", 35)
      Appearance <- "Picture"
   Button "template_test_14" at 0,347 size 130x47; TextOn '6卷绕相关1'; TextOff '6卷绕相关1'
      on Release: ActivateScreenByNumber("Picture", 0); SetTag("ST_HMI_Var_HMI_i32_ZouChe_ZhanJu_ss_1", 0)
      on Press: SetTag("Picture", 36)
      Appearance <- "Picture"
   Button "template_test_15" at 0,413 size 130x47; TextOn '7卷绕相关2'; TextOff '7卷绕相关2'
      on Release: ActivateScreenByNumber("Picture", 0); SetTag("ST_HMI_Var_HMI_i32_ZouChe_ZhanJu_ss_1", 0)
      on Press: SetTag("Picture", 37)
      Appearance <- "Picture"
   Button "template_test_16" at 0,478 size 130x47; TextOn '8存绕相关'; TextOff '8存绕相关'
      on Release: ActivateScreenByNumber("Picture", 0); SetTag("ST_HMI_Var_HMI_i32_ZouChe_ZhanJu_ss_1", 0)
      on Press: SetTag("Picture", 38)
      Appearance <- "Picture"
   Button "template_test_17" at 0,544 size 130x47; TextOn '9自动停止'; TextOff '9自动停止'
      on Release: ActivateScreenByNumber("Picture", 0); SetTag("ST_HMI_Var_HMI_i32_ZouChe_ZhanJu_ss_1", 0)
      on Press: SetTag("Picture", 39)
      Appearance <- "Picture"
   Button "template_test_18" at 0,610 size 130x47; TextOn '10走车相关'; TextOff '10走车相关'
      on Release: ActivateScreenByNumber("Picture", 0); SetTag("ST_HMI_Var_HMI_i32_ZouChe_ZhanJu_ss_1", 0)
      on Press: SetTag("Picture", 40)
      Appearance <- "Picture"
   Button "template_test_19" at 1150,20 size 130x47; TextOn '11生头相关'; TextOff '11生头相关'
      on Release: ActivateScreenByNumber("Picture", 0); SetTag("ST_HMI_Var_HMI_i32_ZouChe_ZhanJu_ss_1", 0)
      on Press: SetTag("Picture", 41)
      Appearance <- "Picture"
   Button "template_test_20" at 1150,85 size 130x47; TextOn '12张力弓整定'; TextOff '12张力弓整定'
      on Release: ActivateScreenByNumber("Picture", 0); SetTag("ST_HMI_Var_HMI_i32_ZouChe_ZhanJu_ss_1", 0)
      on Press: SetTag("Picture", 42)
      Appearance <- "Picture"
   Button "template_test_21" at 1150,150 size 130x47; TextOn '12张力弓整定'; TextOff '13原点设定'
      on Release: ActivateScreenByNumber("Picture", 0); SetTag("ST_HMI_Var_HMI_i32_ZouChe_ZhanJu_ss_1", 0)
      on Press: SetTag("Picture", 43)
      Appearance <- "Picture"
   Button "template_test_22" at 1150,216 size 130x47; TextOn '12张力弓整定'; TextOff '14纱管参数'
      on Release: ActivateScreenByNumber("Picture", 0); SetTag("ST_HMI_Var_HMI_i32_ZouChe_ZhanJu_ss_1", 0)
      on Press: SetTag("Picture", 44)
      Appearance <- "Picture"
   Button "template_test_23" at 160,680 size 160x60; TextOn '工艺'; TextOff '工艺'; PictureOn "settings_1_32×32_反相"; PictureOff "settings_1_32×32"
      on Release: ActivateScreenByNumber("Picture", 0)
      on Press: SetTag("Picture", 2)
      Appearance <- "Picture"
   Button "template_test_24" at 1150,281 size 130x47; TextOn '12张力弓整定'; TextOff '15卷绕经验参数'
      on Release: ActivateScreenByNumber("Picture", 0); SetTag("ST_HMI_Var_HMI_i32_ZouChe_ZhanJu_ss_1", 0)
      on Press: SetTag("Picture", 45)
      Appearance <- "Picture"
   Button "template_test_25" at 1150,347 size 130x47; TextOn '12张力弓整定'; TextOff '16机械参数'
      on Release: ActivateScreenByNumber("Picture", 0); SetTag("ST_HMI_Var_HMI_i32_ZouChe_ZhanJu_ss_1", 0)
      on Press: SetTag("Picture", 46)
      Appearance <- "Picture"
   Button "template_test_26" at 1150,610 size 130x47; TextOn '调试'; TextOff '调试'; PictureOn "图形_18"; PictureOff "图形_18"
      on Release: ActivateScreenByNumber("Picture", 0); SetTag("ST_HMI_Var_HMI_i32_ZouChe_ZhanJu_ss_1", 0)
      on Press: SetTag("Picture", 3)
      Appearance <- "Picture"
   Button "Template_Button_1" at 320,680 size 80x60; TextOff 'Text'; PictureOff "China_1"
      on Click: function_fb9197e8(-1)
   Button "OBJECT_122" at 1200,680 size 80x60; TextOn '响 铃'; TextOff '响 铃 / EXIT'; PictureOn "Gold_bell_100×100_反相"; PictureOff "Gold_bell_100×100"
      on Release: ResetBit("ST_HMI_Var_HMI_bo_XiangLing")
      on Press: SetBit("ST_HMI_Var_HMI_bo_XiangLing")
      Appearance <- "ST_HMI_Var_HMI_bo_XiangLing"

Template "模板_设置" 1280x740
   Button "template_set_1" at 80,680 size 80x60; TextOn '手动画面'; TextOff '手动操作'; PictureOn "manual_5_500×500_反相"; PictureOff "manual_5_500×500"
      on Release: ActivateScreenByNumber("Picture", 0); SetTag("ST_HMI_Var_HMI_i32_ZouChe_ZhanJu_ss_1", 0); function_f23ef4c9()
      on Press: SetTag("Picture", 5)
      Appearance <- "Picture"
   Button "template_set_2" at 720,680 size 80x60; TextOn '报警画面'; TextOff '报 警'; PictureOn "emblem_important_1_200×200_反相"; PictureOff "emblem_important_1_200×200"
      on Release: ActivateScreenByNumber("Picture", 0); SetTag("ST_HMI_Var_HMI_i32_ZouChe_ZhanJu_ss_1", 0); function_f23ef4c9()
      on Press: SetTag("Picture", 6)
      Appearance <- "Picture"
   Button "template_set_5" at 800,680 size 80x60; TextOn '保养提示'; TextOff '保养提示'; PictureOn "baoyang_6_600×600_反相"; PictureOff "baoyang_6_600×600"
      on Release: ActivateScreenByNumber("Picture", 0); SetTag("ST_HMI_Var_HMI_i32_ZouChe_ZhanJu_ss_1", 0); function_f23ef4c9()
      on Press: SetTag("Picture", 8)
      Appearance <- "Picture"
   Button "template_set_7" at 880,680 size 80x60; TextOn '调试画面'; TextOff '调 试'; Authorization "Operate_4"; PictureOff "kdeconnect-tray_100×100"; PictureOn "kdeconnect-tray_100×100_反相"
      on Release: ActivateScreenByNumber("Picture", 0); SetTag("ST_HMI_Var_HMI_i32_ZouChe_ZhanJu_ss_1", 0); function_f23ef4c9()
      on Press: SetTag("Picture", 3)
      Appearance <- "Picture"
   Button "template_set_3" at 0,680 size 80x60; TextOn '手动画面'; TextOff '手动操作'; PictureOff "图形_16"
      on Release: ActivateScreenByNumber("Picture", 0); SetTag("ST_HMI_Var_HMI_i32_ZouChe_ZhanJu_ss_1", 0); function_f23ef4c9()
      on Press: SetTag("Picture", 1)
      Appearance <- "Picture"
   Button "template_set_4" at 1120,680 size 80x60; TextOff '调 试'; TextOn '调试画面'; PictureOn "System_Shutdown_反相_100×100"; PictureOff "System_Shutdown_100×100"; Authorization "Operate_4"
      on Click: function_f23ef4c9()
      on Release: StopRuntime(0); function_f23ef4c9(); SetTag("ST_HMI_Var_HMI_i32_ZouChe_ZhanJu_ss_1", 0)
   Button "template_set_6" at 1040,680 size 80x60; TextOff 'Text'; TextOn '调试画面'; PictureOn "computer_laptop_100×100_反相"; PictureOff "computer_laptop_100×100"; Authorization "Operate_4"
      on Click: function_f23ef4c9()
      on Release: function_f34a74f3(); function_f23ef4c9(); SetTag("ST_HMI_Var_HMI_i32_ZouChe_ZhanJu_ss_1", 0)
   Button "template_set_8" at 960,680 size 80x60; TextOff 'Text'; TextOn '调试画面'; PictureOn "similarartists_amarok_100×100_反相"; PictureOff "similarartists_amarok_100×100"; Authorization "Operate_4"
      on Release: ActivateScreenByNumber("Picture", 0); SetTag("ST_HMI_Var_HMI_i32_ZouChe_ZhanJu_ss_1", 0); function_f23ef4c9()
      on Press: SetTag("Picture", 7)
      Appearance <- "Picture"
   Button "template_set_23" at 160,680 size 160x60; TextOn '工艺'; TextOff '工艺'; PictureOn "settings_1_32×32_反相"; PictureOff "settings_1_32×32"
      on Release: ActivateScreenByNumber("Picture", 0); SetTag("ST_HMI_Var_HMI_i32_ZouChe_ZhanJu_ss_1", 0); function_f23ef4c9()
      on Press: SetTag("Picture", 2)
      Appearance <- "Picture"
   Button "template_set_10" at 1150,24 size 130x47; TextOn '车况设定'; TextOff '车况设定'; Authorization "Operate_5"
      on Release: ActivateScreenByNumber("Picture", 0)
      on Press: SetTag("Picture", 21)
      Appearance <- "Picture"
   Button "template_set_11" at 1150,107 size 130x47; TextOn '纱穗参数设定'; TextOff '纱穗参数'; Authorization "Operate_5"
      on Release: ActivateScreenByNumber("Picture", 0)
      on Press: SetTag("Picture", 22)
      Appearance <- "Picture"
   Button "template_set_12" at 1150,191 size 130x47; TextOn '退绕设定'; TextOff '退绕设定'; Authorization "Operate_5"
      on Release: ActivateScreenByNumber("Picture", 0)
      on Press: SetTag("Picture", 23)
      Appearance <- "Picture"
   Button "template_set_13" at 1150,358 size 130x47; TextOn '退绕设定'; TextOff '牵伸曲线'
      on Release: ActivateScreenByNumber("Picture", 0)
      on Press: SetTag("Picture", 25)
      Appearance <- "Picture"
   Button "按钮_1" at 1150,275 size 130x47; TextOff '牵伸调整'; Authorization "Operate_5"
      on Release: ActivateScreenByNumber("Picture", 0)
      on Press: SetTag("Picture", 24)
      Appearance <- "Picture"
   Button "template_set_26" at 1150,610 size 130x47; TextOn '设置'; TextOff '设置'; PictureOn "图形_17"; PictureOff "图形_17"
      on Release: ActivateScreenByNumber("Picture", 0); function_f23ef4c9()
      on Press: SetTag("Picture", 2)
      Appearance <- "Picture"
   TextField "模板_文本域_2" at 320,680 size 400x60; Text '苏州友联纺工装备科技股份有限公司'
   Button "template_set_9" at 1150,442 size 130x47; TextOn '退绕设定'; TextOff '分段捻缩'; Authorization "Operate_5"
      on Release: ActivateScreenByNumber("Picture", 0)
      on Press: SetTag("Picture", 26)
      Appearance <- "Picture"
   Button "template_set_14" at 1150,526 size 130x47; TextOn '退绕设定'; TextOff '包芯纱'; Authorization "Operate_5"
      on Release: ActivateScreenByNumber("Picture", 0)
      on Press: SetTag("Picture", 27)
      Appearance <- "Picture"
   Button "OBJECT_122" at 1200,680 size 80x60; TextOn '响 铃'; TextOff '响 铃 / EXIT'; PictureOn "Gold_bell_100×100_反相"; PictureOff "Gold_bell_100×100"
      on Release: ResetBit("ST_HMI_Var_HMI_bo_XiangLing")
      on Press: SetBit("ST_HMI_Var_HMI_bo_XiangLing")
      Appearance <- "ST_HMI_Var_HMI_bo_XiangLing"

screen "监控画面" 1280x740, template "模板_根"
   IOField "IO Field_3" at 48,24 size 128x42; FormatPattern 99.999
      ProcessValue <- "ST_Real_Monitoring_HMI_r64_Real_QianShen_WuNian"
   IOField "IO Field_1" at 48,80 size 128x42; FormatPattern 99.999
      ProcessValue <- "ST_HMI_Var_HMI_r64QianShen_All_real"
   IOField "IO Field_2" at 48,144 size 128x42; FormatPattern 9999.99
      ProcessValue <- "ST_Real_Monitoring_HMI_r64Axis_ZouChe_Position_JiZhong_QianShen_Start"
   IOField "IO Field_4" at 48,200 size 128x42; FormatPattern 9999
      ProcessValue <- "ST_Real_Monitoring_HMI_r64_NianDu_JiZhong_QianShen_Start"
   IOField "IO Field_5" at 48,264 size 128x42; FormatPattern 9999.99
      ProcessValue <- "ST_Real_Monitoring_HMI_r64Axis_ZouChe_Position_LuoLa_Stop"
   IOField "IO Field_6" at 48,320 size 128x42; FormatPattern 9999
      ProcessValue <- "ST_Real_Monitoring_HMI_r64_NianDu_LuoLa_Stop"
   IOField "IO Field_7" at 48,384 size 128x42; FormatPattern 9999
      ProcessValue <- "ST_HMI_Var_HMI_r64NianDu_actual"
   IOField "IO Field_8" at 48,440 size 128x42; FormatPattern 9999.99
      ProcessValue <- "ST_Real_Monitoring_HMI_r64Axis_ZouChe_Position_YiNian_DaoDa"
   IOField "IO Field_10" at 588,24 size 128x42; FormatPattern 99.999
      ProcessValue <- "ST_Convert_ReadParameters_g_r64_SERVO_03_ZouChe_35_Motor_temperature_real"
   IOField "IO Field_11" at 588,81 size 128x42; FormatPattern 999.99
      ProcessValue <- "ST_Convert_ReadParameters_g_r64_SERVO_04_ZhangLi_35_Motor_temperature_real"
   IOField "IO Field_12" at 588,138 size 128x42; FormatPattern 999.99
      ProcessValue <- "ST_Convert_ReadParameters_g_r64_SERVO_05_ChengXing_35_Motor_temperature_real"
   IOField "IO Field_13" at 588,195 size 128x42; FormatPattern 999.99
      ProcessValue <- "ST_Convert_ReadParameters_g_r64_SERVO_06_GunTong_35_Motor_temperature_real"
   IOField "IO Field_14" at 588,252 size 128x42; FormatPattern 999.99
      ProcessValue <- "ST_Convert_ReadParameters_g_r64_SERVO_08_LuoLa_35_Motor_temperature_real"
   IOField "IO Field_15" at 588,309 size 128x42; FormatPattern 999.99
      ProcessValue <- "ST_Convert_ReadParameters_g_r64_SERVO_07_DingZi_35_Motor_temperature_real"
   IOField "IO Field_17" at 588,366 size 128x42; FormatPattern 999.99
      ProcessValue <- "ST_Convert_ReadParameters_g_r64_SERVO_03_ZouChe_37_4_Power_unit_temperatures_Interior_of_power_unit_real"
   IOField "IO Field_18" at 588,423 size 128x42; FormatPattern 999.99
      ProcessValue <- "ST_Convert_ReadParameters_g_r64_SERVO_05_ChengXing_37_4_Power_unit_temperatures_Interior_of_power_unit_real"
   IOField "IO Field_19" at 588,480 size 128x42; FormatPattern 999.99
      ProcessValue <- "ST_Convert_ReadParameters_g_r64_SERVO_07_DingZi_37_4_Power_unit_temperatures_Interior_of_power_unit_real"
   IOField "IO Field_20" at 588,538 size 128x42; FormatPattern 999.99
      ProcessValue <- "ST_Convert_ReadParameters_g_r64_SERVO_08_LuoLa_37_4_Power_unit_temperatures_Interior_of_power_unit_real"
   TextField "Text Field_40" at 191,24 size 352x42; Text '实时无捻牵伸 / 番手: / 실 번수'
   TextField "Text Field_1" at 193,80 size 352x42; Text '实时总牵伸 / 番手: / 실 번수'
   TextField "Text Field_2" at 194,144 size 352x42; Text '集中牵伸开始时的走车位置 / 番手: / 실 번수'
   TextField "Text Field_3" at 193,200 size 352x42; Text '集中牵伸开始时的捻度 / 番手: / 실 번수'
   TextField "Text Field_4" at 195,264 size 352x42; Text '罗拉停止时的走车位置 / 番手: / 실 번수'
   TextField "Text Field_5" at 194,320 size 352x42; Text '罗拉停止时的捻度 / 番手: / 실 번수'
   TextField "Text Field_6" at 194,384 size 352x42; Text '实际捻度 / 番手: / 실 번수'
   TextField "Text Field_7" at 193,440 size 352x42; Text '锭子加速到第一个峰值时的走车位置 / 番手: / 실 번수'
   TextField "Text Field_9" at 732,24 size 352x42; Text '走车电机实时温度（℃） / 番手: / 실 번수'
   TextField "Text Field_10" at 732,81 size 352x42; Text '张力电机实时温度（℃） / 番手: / 실 번수'
   TextField "Text Field_11" at 732,138 size 352x42; Text '成形电机实时温度（℃） / 番手: / 실 번수'
   TextField "Text Field_12" at 732,195 size 352x42; Text '滚筒电机实时温度（℃） / 番手: / 실 번수'
   TextField "Text Field_13" at 732,252 size 352x42; Text '罗拉电机实时温度（℃） / 番手: / 실 번수'
   TextField "Text Field_14" at 732,309 size 352x42; Text '锭子电机实时温度（℃） / 番手: / 실 번수'
   TextField "Text Field_16" at 732,366 size 352x42; Text '走车张力驱动器实时温度（℃） / 番手: / 실 번수'
   TextField "Text Field_17" at 732,423 size 352x42; Text '成形滚筒驱动器实时温度（℃） / 番手: / 실 번수'
   TextField "Text Field_18" at 732,480 size 352x42; Text '锭子驱动器实时温度（℃） / 番手: / 실 번수'
   TextField "Text Field_19" at 732,538 size 352x42; Text '罗拉驱动器实时温度（℃） / 番手: / 실 번수'
   Button "HmiScreenItemData_6" at 1150,396 size 130x47; TextOn '12张力弓整定'; TextOff '返回'
      on Release: ActivateScreenByNumber("Picture", 0); SetTag("ST_HMI_Var_HMI_i32_ZouChe_ZhanJu_ss_1", 0)
      on Press: SetTag("Picture", 6)

